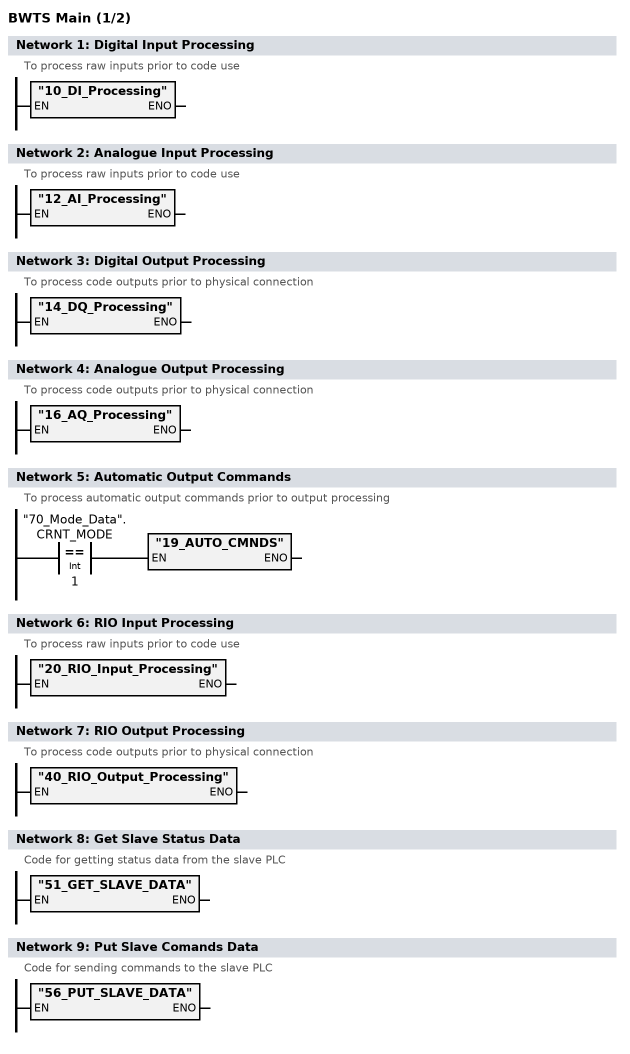
   RUNG wire#powerrail
      "10_DI_Processing"()
   END_RUNG
   // the same network as SCL:
   "10_DI_Processing"();
END_REGION

REGION Network 2: Analogue Input Processing
   // To process raw inputs prior to code use
   RUNG wire#powerrail
      "12_AI_Processing"()
   END_RUNG
   // the same network as SCL:
   "12_AI_Processing"();
END_REGION

REGION Network 3: Digital Output Processing
   // To process code outputs prior to physical connection
   RUNG wire#powerrail
      "14_DQ_Processing"()
   END_RUNG
   // the same network as SCL:
   "14_DQ_Processing"();
END_REGION

REGION Network 4: Analogue Output Processing
   // To process code outputs prior to physical connection
   RUNG wire#powerrail
      "16_AQ_Processing"()
   END_RUNG
   // the same network as SCL:
   "16_AQ_Processing"();
END_REGION

REGION Network 5: Automatic Output Commands
   // To process automatic output commands prior to output processing
   RUNG wire#powerrail
      { S7_Templates := "SrcType := Int" } EQ_Contact(in1 := "70_Mode_Data".CRNT_MODE, in2 := 1)
      "19_AUTO_CMNDS"()
   END_RUNG
   // the same network as SCL:
   IF "70_Mode_Data".CRNT_MODE = 1 THEN "19_AUTO_CMNDS"(); END_IF;
END_REGION

REGION Network 6: RIO Input Processing
   // To process raw inputs prior to code use
   RUNG wire#powerrail
      "20_RIO_Input_Processing"()
   END_RUNG
   // the same network as SCL:
   "20_RIO_Input_Processing"();
END_REGION

REGION Network 7: RIO Output Processing
   // To process code outputs prior to physical connection
   RUNG wire#powerrail
      "40_RIO_Output_Processing"()
   END_RUNG
   // the same network as SCL:
   "40_RIO_Output_Processing"();
END_REGION

REGION Network 8: Get Slave Status Data
   // Code for getting status data from the slave PLC
   RUNG wire#powerrail
      "51_GET_SLAVE_DATA"()
   END_RUNG
   // the same network as SCL:
   "51_GET_SLAVE_DATA"();
END_REGION

REGION Network 9: Put Slave Comands Data
   // Code for sending commands to the slave PLC
   RUNG wire#powerrail
      "56_PUT_SLAVE_DATA"()
   END_RUNG
   // the same network as SCL:
   "56_PUT_SLAVE_DATA"();
END_REGION

REGION Network 10: Communications Heart Beat
   // Code for communications heart beat bit
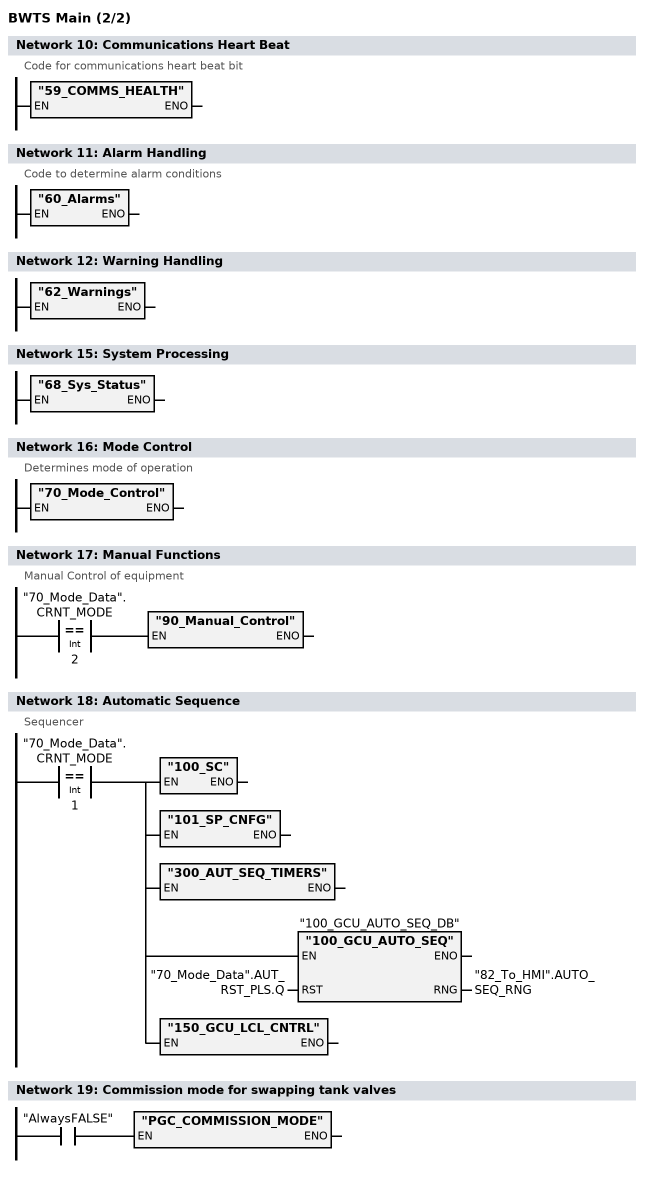
   RUNG wire#powerrail
      "59_COMMS_HEALTH"()
   END_RUNG
   // the same network as SCL:
   "59_COMMS_HEALTH"();
END_REGION

REGION Network 11: Alarm Handling
   // Code to determine alarm conditions
   RUNG wire#powerrail
      "60_Alarms"()
   END_RUNG
   // the same network as SCL:
   "60_Alarms"();
END_REGION

REGION Network 12: Warning Handling
   RUNG wire#powerrail
      "62_Warnings"()
   END_RUNG
   // the same network as SCL:
   "62_Warnings"();
END_REGION

REGION Network 13: Message Handling
   // Handles messaging
END_REGION

REGION Network 14: Event Handling
   // Records event data
END_REGION

REGION Network 15: System Processing
   RUNG wire#powerrail
      "68_Sys_Status"()
   END_RUNG
   // the same network as SCL:
   "68_Sys_Status"();
END_REGION

REGION Network 16: Mode Control
   // Determines mode of operation
   RUNG wire#powerrail
      "70_Mode_Control"()
   END_RUNG
   // the same network as SCL:
   "70_Mode_Control"();
END_REGION

REGION Network 17: Manual Functions
   // Manual Control of equipment
   RUNG wire#powerrail
      { S7_Templates := "SrcType := Int" } EQ_Contact(in1 := "70_Mode_Data".CRNT_MODE, in2 := 2)
      "90_Manual_Control"()
   END_RUNG
   // the same network as SCL:
   IF "70_Mode_Data".CRNT_MODE = 2 THEN "90_Manual_Control"(); END_IF;
END_REGION

REGION Network 18: Automatic Sequence
   // Sequencer
   RUNG wire#powerrail
      { S7_Templates := "SrcType := Int" } EQ_Contact(in1 := "70_Mode_Data".CRNT_MODE, in2 := 1)
      wire#w1
      "100_SC"()
   END_RUNG
   RUNG wire#w1
      "101_SP_CNFG"()
   END_RUNG
   RUNG wire#w1
      "300_AUT_SEQ_TIMERS"()
   END_RUNG
   RUNG wire#w1
      "100_GCU_AUTO_SEQ_DB"(RST := "70_Mode_Data".AUT_RST_PLS.Q, RNG => "82_To_HMI".AUTO_SEQ_RNG)
   END_RUNG
   RUNG wire#w1
      "150_GCU_LCL_CNTRL"()
   END_RUNG
   // the same network as SCL:
   #_w1 := "70_Mode_Data".CRNT_MODE = 1;
   IF #_w1 THEN
       "100_SC"();
       "101_SP_CNFG"();
       "300_AUT_SEQ_TIMERS"();
       "100_GCU_AUTO_SEQ_DB"(RST := "70_Mode_Data".AUT_RST_PLS.Q, RNG => "82_To_HMI".AUTO_SEQ_RNG);   // "100_GCU_AUTO_SEQ"
       "150_GCU_LCL_CNTRL"();
   END_IF;
END_REGION

REGION Network 19: Commission mode for swapping tank valves
   RUNG wire#powerrail
      Contact( "AlwaysFALSE" )
      "PGC_COMMISSION_MODE"()
   END_RUNG
   // the same network as SCL:
   IF "AlwaysFALSE" THEN "PGC_COMMISSION_MODE"(); END_IF;
END_REGION
END_ORGANIZATION_BLOCK

// folder: 10 - 19 IO & Processing

FUNCTION "10_DI_Processing" : Void   // FC10, LAD
TITLE = Digital Input Processing
{ S7_Optimized_Access := 'TRUE' }
AUTHOR : JRS
VERSION : 0.1
// To process raw inputs prior to code use
BEGIN

REGION Network 1: I136.0 - Spare Input
   // True = N/A, False = N/A
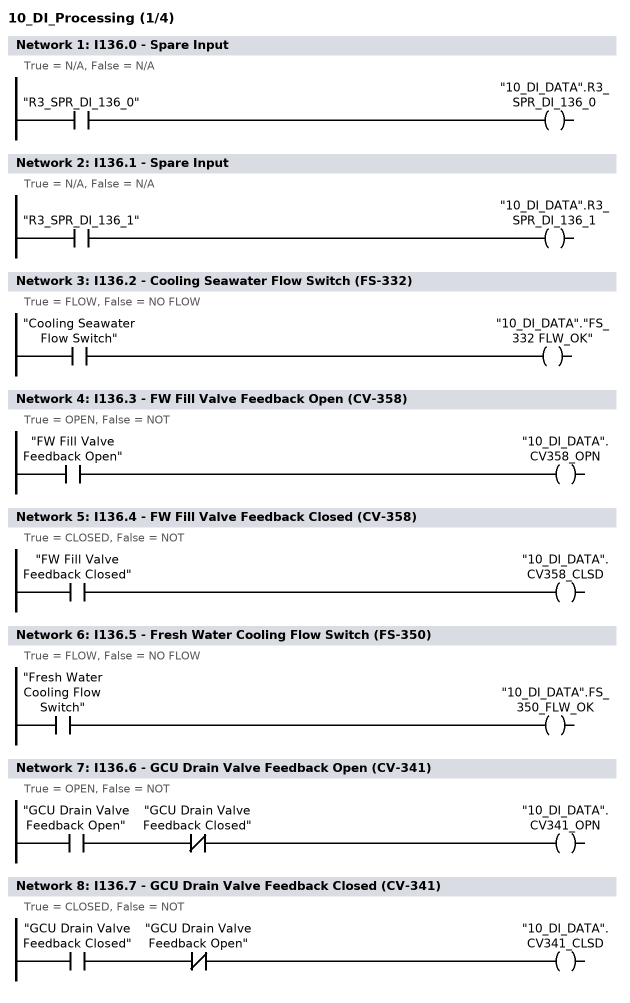
   RUNG wire#powerrail
      Contact( "R3_SPR_DI_136_0" )
      Coil( "10_DI_DATA".R3_SPR_DI_136_0 )
   END_RUNG
   // the same network as SCL:
   "10_DI_DATA".R3_SPR_DI_136_0 := "R3_SPR_DI_136_0";
END_REGION

REGION Network 2: I136.1 - Spare Input
   // True = N/A, False = N/A
   RUNG wire#powerrail
      Contact( "R3_SPR_DI_136_1" )
      Coil( "10_DI_DATA".R3_SPR_DI_136_1 )
   END_RUNG
   // the same network as SCL:
   "10_DI_DATA".R3_SPR_DI_136_1 := "R3_SPR_DI_136_1";
END_REGION

REGION Network 3: I136.2 - Cooling Seawater Flow Switch (FS-332)
   // True = FLOW, False = NO FLOW
   RUNG wire#powerrail
      Contact( "Cooling Seawater Flow Switch" )
      Coil( "10_DI_DATA"."FS_332 FLW_OK" )
   END_RUNG
   // the same network as SCL:
   "10_DI_DATA"."FS_332 FLW_OK" := "Cooling Seawater Flow Switch";
END_REGION

REGION Network 4: I136.3 - FW Fill Valve Feedback Open (CV-358)
   // True = OPEN, False = NOT
   RUNG wire#powerrail
      Contact( "FW Fill Valve Feedback Open" )
      Coil( "10_DI_DATA".CV358_OPN )
   END_RUNG
   // the same network as SCL:
   "10_DI_DATA".CV358_OPN := "FW Fill Valve Feedback Open";
END_REGION

REGION Network 5: I136.4 - FW Fill Valve Feedback Closed (CV-358)
   // True = CLOSED, False = NOT
   RUNG wire#powerrail
      Contact( "FW Fill Valve Feedback Closed" )
      Coil( "10_DI_DATA".CV358_CLSD )
   END_RUNG
   // the same network as SCL:
   "10_DI_DATA".CV358_CLSD := "FW Fill Valve Feedback Closed";
END_REGION

REGION Network 6: I136.5 - Fresh Water Cooling Flow Switch (FS-350)
   // True = FLOW, False = NO FLOW
   RUNG wire#powerrail
      Contact( "Fresh Water Cooling Flow Switch" )
      Coil( "10_DI_DATA".FS_350_FLW_OK )
   END_RUNG
   // the same network as SCL:
   "10_DI_DATA".FS_350_FLW_OK := "Fresh Water Cooling Flow Switch";
END_REGION

REGION Network 7: I136.6 - GCU Drain Valve Feedback Open (CV-341)
   // True = OPEN, False = NOT
   RUNG wire#powerrail
      Contact( "GCU Drain Valve Feedback Open" )
      I_Contact( "GCU Drain Valve Feedback Closed" )
      Coil( "10_DI_DATA".CV341_OPN )
   END_RUNG
   // the same network as SCL:
   "10_DI_DATA".CV341_OPN := "GCU Drain Valve Feedback Open" AND NOT "GCU Drain Valve Feedback Closed";
END_REGION

REGION Network 8: I136.7 - GCU Drain Valve Feedback Closed (CV-341)
   // True = CLOSED, False = NOT
   RUNG wire#powerrail
      Contact( "GCU Drain Valve Feedback Closed" )
      I_Contact( "GCU Drain Valve Feedback Open" )
      Coil( "10_DI_DATA".CV341_CLSD )
   END_RUNG
   // the same network as SCL:
   "10_DI_DATA".CV341_CLSD := "GCU Drain Valve Feedback Closed" AND NOT "GCU Drain Valve Feedback Open";
END_REGION

REGION Network 9: I137.0 - Gas to Deck Valve Feedback Open (CV-406)
   // True = OPEN, False = NOT
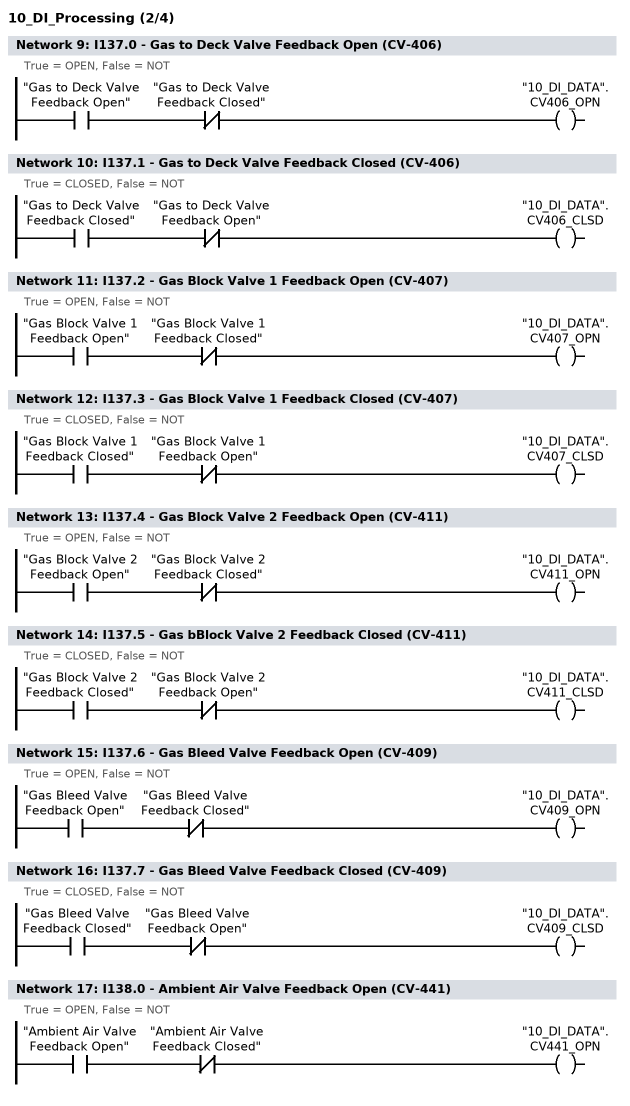
   RUNG wire#powerrail
      Contact( "Gas to Deck Valve Feedback Open" )
      I_Contact( "Gas to Deck Valve Feedback Closed" )
      Coil( "10_DI_DATA".CV406_OPN )
   END_RUNG
   // the same network as SCL:
   "10_DI_DATA".CV406_OPN := "Gas to Deck Valve Feedback Open" AND NOT "Gas to Deck Valve Feedback Closed";
END_REGION

REGION Network 10: I137.1 - Gas to Deck Valve Feedback Closed (CV-406)
   // True = CLOSED, False = NOT
   RUNG wire#powerrail
      Contact( "Gas to Deck Valve Feedback Closed" )
      I_Contact( "Gas to Deck Valve Feedback Open" )
      Coil( "10_DI_DATA".CV406_CLSD )
   END_RUNG
   // the same network as SCL:
   "10_DI_DATA".CV406_CLSD := "Gas to Deck Valve Feedback Closed" AND NOT "Gas to Deck Valve Feedback Open";
END_REGION

REGION Network 11: I137.2 - Gas Block Valve 1 Feedback Open (CV-407)
   // True = OPEN, False = NOT
   RUNG wire#powerrail
      Contact( "Gas Block Valve 1 Feedback Open" )
      I_Contact( "Gas Block Valve 1 Feedback Closed" )
      Coil( "10_DI_DATA".CV407_OPN )
   END_RUNG
   // the same network as SCL:
   "10_DI_DATA".CV407_OPN := "Gas Block Valve 1 Feedback Open" AND NOT "Gas Block Valve 1 Feedback Closed";
END_REGION

REGION Network 12: I137.3 - Gas Block Valve 1 Feedback Closed (CV-407)
   // True = CLOSED, False = NOT
   RUNG wire#powerrail
      Contact( "Gas Block Valve 1 Feedback Closed" )
      I_Contact( "Gas Block Valve 1 Feedback Open" )
      Coil( "10_DI_DATA".CV407_CLSD )
   END_RUNG
   // the same network as SCL:
   "10_DI_DATA".CV407_CLSD := "Gas Block Valve 1 Feedback Closed" AND NOT "Gas Block Valve 1 Feedback Open";
END_REGION

REGION Network 13: I137.4 - Gas Block Valve 2 Feedback Open (CV-411)
   // True = OPEN, False = NOT
   RUNG wire#powerrail
      Contact( "Gas Block Valve 2 Feedback Open" )
      I_Contact( "Gas Block Valve 2 Feedback Closed" )
      Coil( "10_DI_DATA".CV411_OPN )
   END_RUNG
   // the same network as SCL:
   "10_DI_DATA".CV411_OPN := "Gas Block Valve 2 Feedback Open" AND NOT "Gas Block Valve 2 Feedback Closed";
END_REGION

REGION Network 14: I137.5 - Gas bBlock Valve 2 Feedback Closed (CV-411)
   // True = CLOSED, False = NOT
   RUNG wire#powerrail
      Contact( "Gas Block Valve 2 Feedback Closed" )
      I_Contact( "Gas Block Valve 2 Feedback Open" )
      Coil( "10_DI_DATA".CV411_CLSD )
   END_RUNG
   // the same network as SCL:
   "10_DI_DATA".CV411_CLSD := "Gas Block Valve 2 Feedback Closed" AND NOT "Gas Block Valve 2 Feedback Open";
END_REGION

REGION Network 15: I137.6 - Gas Bleed Valve Feedback Open (CV-409)
   // True = OPEN, False = NOT
   RUNG wire#powerrail
      Contact( "Gas Bleed Valve Feedback Open" )
      I_Contact( "Gas Bleed Valve Feedback Closed" )
      Coil( "10_DI_DATA".CV409_OPN )
   END_RUNG
   // the same network as SCL:
   "10_DI_DATA".CV409_OPN := "Gas Bleed Valve Feedback Open" AND NOT "Gas Bleed Valve Feedback Closed";
END_REGION

REGION Network 16: I137.7 - Gas Bleed Valve Feedback Closed (CV-409)
   // True = CLOSED, False = NOT
   RUNG wire#powerrail
      Contact( "Gas Bleed Valve Feedback Closed" )
      I_Contact( "Gas Bleed Valve Feedback Open" )
      Coil( "10_DI_DATA".CV409_CLSD )
   END_RUNG
   // the same network as SCL:
   "10_DI_DATA".CV409_CLSD := "Gas Bleed Valve Feedback Closed" AND NOT "Gas Bleed Valve Feedback Open";
END_REGION

REGION Network 17: I138.0 - Ambient Air Valve Feedback Open (CV-441)
   // True = OPEN, False = NOT
   RUNG wire#powerrail
      Contact( "Ambient Air Valve Feedback Open" )
      I_Contact( "Ambient Air Valve Feedback Closed" )
      Coil( "10_DI_DATA".CV441_OPN )
   END_RUNG
   // the same network as SCL:
   "10_DI_DATA".CV441_OPN := "Ambient Air Valve Feedback Open" AND NOT "Ambient Air Valve Feedback Closed";
END_REGION

REGION Network 18: I138.1 - Ambient Air Valve Feedback Closed (CV-441)
   // True = CLOSED, False = NOT
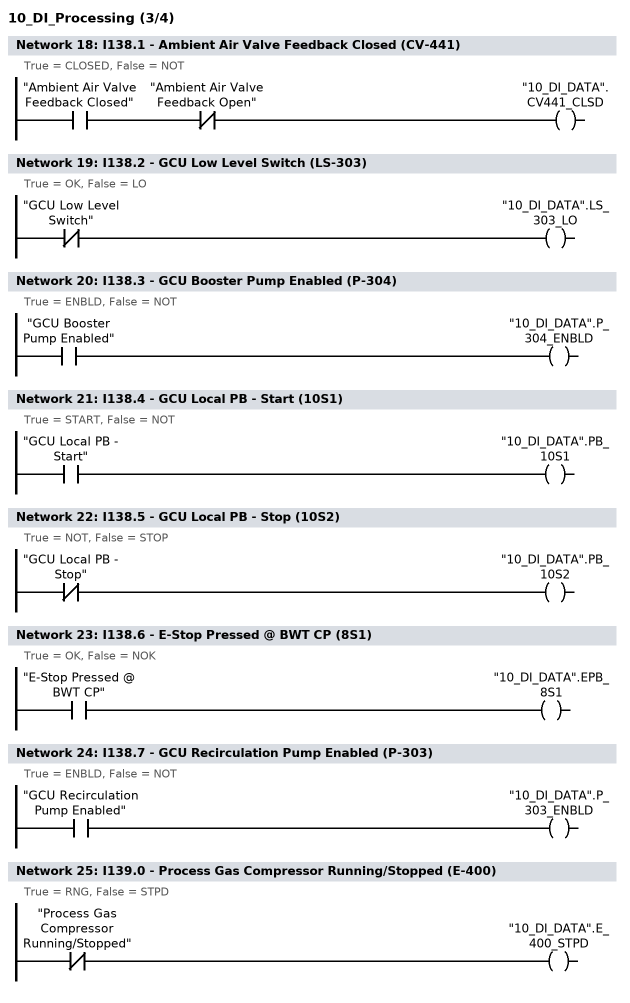
   RUNG wire#powerrail
      Contact( "Ambient Air Valve Feedback Closed" )
      I_Contact( "Ambient Air Valve Feedback Open" )
      Coil( "10_DI_DATA".CV441_CLSD )
   END_RUNG
   // the same network as SCL:
   "10_DI_DATA".CV441_CLSD := "Ambient Air Valve Feedback Closed" AND NOT "Ambient Air Valve Feedback Open";
END_REGION

REGION Network 19: I138.2 - GCU Low Level Switch (LS-303)
   // True = OK, False = LO
   RUNG wire#powerrail
      I_Contact( "GCU Low Level Switch" )
      Coil( "10_DI_DATA".LS_303_LO )
   END_RUNG
   // the same network as SCL:
   "10_DI_DATA".LS_303_LO := NOT "GCU Low Level Switch";
END_REGION

REGION Network 20: I138.3 - GCU Booster Pump Enabled (P-304)
   // True = ENBLD, False = NOT
   RUNG wire#powerrail
      Contact( "GCU Booster Pump Enabled" )
      Coil( "10_DI_DATA".P_304_ENBLD )
   END_RUNG
   // the same network as SCL:
   "10_DI_DATA".P_304_ENBLD := "GCU Booster Pump Enabled";
END_REGION

REGION Network 21: I138.4 - GCU Local PB - Start (10S1)
   // True = START, False = NOT
   RUNG wire#powerrail
      Contact( "GCU Local PB - Start" )
      Coil( "10_DI_DATA".PB_10S1 )
   END_RUNG
   // the same network as SCL:
   "10_DI_DATA".PB_10S1 := "GCU Local PB - Start";
END_REGION

REGION Network 22: I138.5 - GCU Local PB - Stop (10S2)
   // True = NOT, False = STOP
   RUNG wire#powerrail
      I_Contact( "GCU Local PB - Stop" )
      Coil( "10_DI_DATA".PB_10S2 )
   END_RUNG
   // the same network as SCL:
   "10_DI_DATA".PB_10S2 := NOT "GCU Local PB - Stop";
END_REGION

REGION Network 23: I138.6 - E-Stop Pressed @ BWT CP (8S1)
   // True = OK, False = NOK
   RUNG wire#powerrail
      Contact( "E-Stop Pressed @ BWT CP" )
      Coil( "10_DI_DATA".EPB_8S1 )
   END_RUNG
   // the same network as SCL:
   "10_DI_DATA".EPB_8S1 := "E-Stop Pressed @ BWT CP";
END_REGION

REGION Network 24: I138.7 - GCU Recirculation Pump Enabled (P-303)
   // True = ENBLD, False = NOT
   RUNG wire#powerrail
      Contact( "GCU Recirculation Pump Enabled" )
      Coil( "10_DI_DATA".P_303_ENBLD )
   END_RUNG
   // the same network as SCL:
   "10_DI_DATA".P_303_ENBLD := "GCU Recirculation Pump Enabled";
END_REGION

REGION Network 25: I139.0 - Process Gas Compressor Running/Stopped (E-400)
   // True = RNG, False = STPD
   RUNG wire#powerrail
      I_Contact( "Process Gas Compressor Running/Stopped" )
      Coil( "10_DI_DATA".E_400_STPD )
   END_RUNG
   // the same network as SCL:
   "10_DI_DATA".E_400_STPD := NOT "Process Gas Compressor Running/Stopped";
END_REGION

REGION Network 26: I139.1 - Process Gas Compressor Tripped/Shutdown (E-400)
   // True = NOK, False = OK
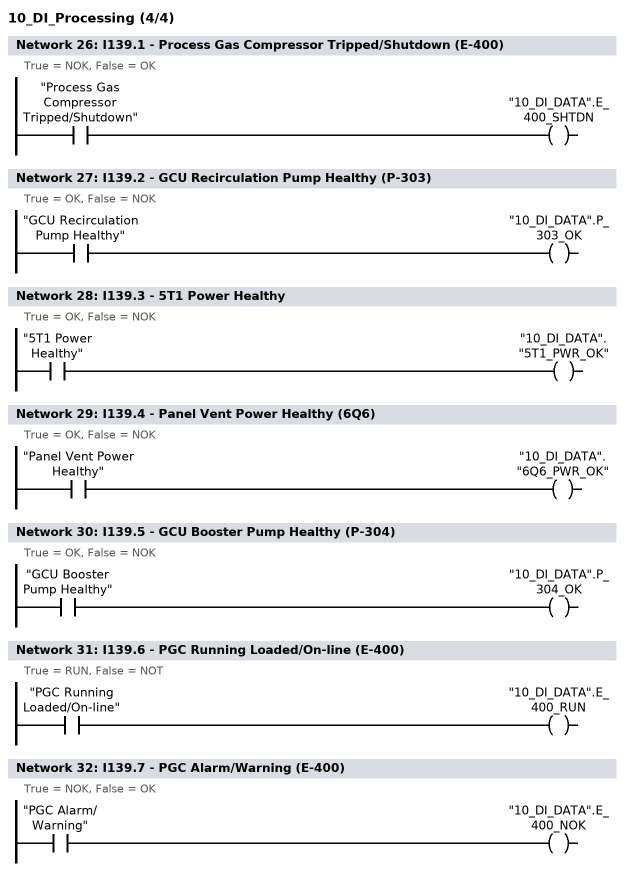
   RUNG wire#powerrail
      Contact( "Process Gas Compressor Tripped/Shutdown" )
      Coil( "10_DI_DATA".E_400_SHTDN )
   END_RUNG
   // the same network as SCL:
   "10_DI_DATA".E_400_SHTDN := "Process Gas Compressor Tripped/Shutdown";
END_REGION

REGION Network 27: I139.2 - GCU Recirculation Pump Healthy (P-303)
   // True = OK, False = NOK
   RUNG wire#powerrail
      Contact( "GCU Recirculation Pump Healthy" )
      Coil( "10_DI_DATA".P_303_OK )
   END_RUNG
   // the same network as SCL:
   "10_DI_DATA".P_303_OK := "GCU Recirculation Pump Healthy";
END_REGION

REGION Network 28: I139.3 - 5T1 Power Healthy
   // True = OK, False = NOK
   RUNG wire#powerrail
      Contact( "5T1 Power Healthy" )
      Coil( "10_DI_DATA"."5T1_PWR_OK" )
   END_RUNG
   // the same network as SCL:
   "10_DI_DATA"."5T1_PWR_OK" := "5T1 Power Healthy";
END_REGION

REGION Network 29: I139.4 - Panel Vent Power Healthy (6Q6)
   // True = OK, False = NOK
   RUNG wire#powerrail
      Contact( "Panel Vent Power Healthy" )
      Coil( "10_DI_DATA"."6Q6_PWR_OK" )
   END_RUNG
   // the same network as SCL:
   "10_DI_DATA"."6Q6_PWR_OK" := "Panel Vent Power Healthy";
END_REGION

REGION Network 30: I139.5 - GCU Booster Pump Healthy (P-304)
   // True = OK, False = NOK
   RUNG wire#powerrail
      Contact( "GCU Booster Pump Healthy" )
      Coil( "10_DI_DATA".P_304_OK )
   END_RUNG
   // the same network as SCL:
   "10_DI_DATA".P_304_OK := "GCU Booster Pump Healthy";
END_REGION

REGION Network 31: I139.6 - PGC Running Loaded/On-line (E-400)
   // True = RUN, False = NOT
   RUNG wire#powerrail
      Contact( "PGC Running Loaded/On-line" )
      Coil( "10_DI_DATA".E_400_RUN )
   END_RUNG
   // the same network as SCL:
   "10_DI_DATA".E_400_RUN := "PGC Running Loaded/On-line";
END_REGION

REGION Network 32: I139.7 - PGC Alarm/Warning (E-400)
   // True = NOK, False = OK
   RUNG wire#powerrail
      Contact( "PGC Alarm/Warning" )
      Coil( "10_DI_DATA".E_400_NOK )
   END_RUNG
   // the same network as SCL:
   "10_DI_DATA".E_400_NOK := "PGC Alarm/Warning";
END_REGION
END_FUNCTION

FUNCTION "12_AI_Processing" : Void   // FC12, LAD
TITLE = Analogue Input Processing
{ S7_Optimized_Access := 'TRUE' }
AUTHOR : JRS
VERSION : 0.1
// To process raw inputs prior to code use
BEGIN

REGION Network 1: IW800 - GCU Level (LIT-304)
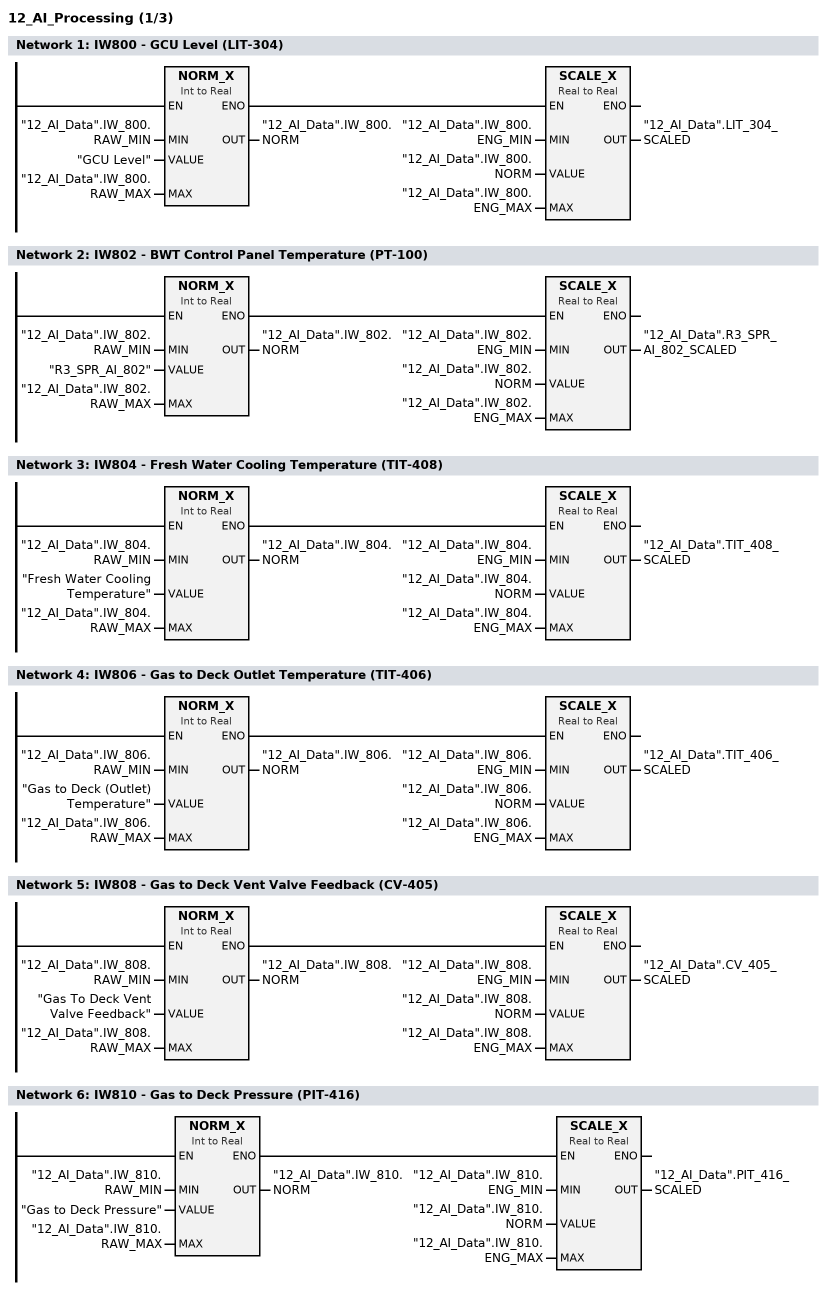
   RUNG wire#powerrail
      { S7_Templates := "[SrcType := Int, DestType := Real]" } Normalize(min := "12_AI_Data".IW_800.RAW_MIN, value := "GCU Level", max := "12_AI_Data".IW_800.RAW_MAX, out => "12_AI_Data".IW_800.NORM)
      { S7_Templates := "[SrcType := Real, DestType := Real]" } Scale(min := "12_AI_Data".IW_800.ENG_MIN, value := "12_AI_Data".IW_800.NORM, max := "12_AI_Data".IW_800.ENG_MAX, out => "12_AI_Data".LIT_304_SCALED)
   END_RUNG
   // the same network as SCL:
   "12_AI_Data".IW_800.NORM := NORM_X(MIN := "12_AI_Data".IW_800.RAW_MIN, VALUE := "GCU Level", MAX := "12_AI_Data".IW_800.RAW_MAX);
   "12_AI_Data".LIT_304_SCALED := SCALE_X(MIN := "12_AI_Data".IW_800.ENG_MIN, VALUE := "12_AI_Data".IW_800.NORM, MAX := "12_AI_Data".IW_800.ENG_MAX);
END_REGION

REGION Network 2: IW802 - BWT Control Panel Temperature (PT-100)
   RUNG wire#powerrail
      { S7_Templates := "[SrcType := Int, DestType := Real]" } Normalize(min := "12_AI_Data".IW_802.RAW_MIN, value := "R3_SPR_AI_802", max := "12_AI_Data".IW_802.RAW_MAX, out => "12_AI_Data".IW_802.NORM)
      { S7_Templates := "[SrcType := Real, DestType := Real]" } Scale(min := "12_AI_Data".IW_802.ENG_MIN, value := "12_AI_Data".IW_802.NORM, max := "12_AI_Data".IW_802.ENG_MAX, out => "12_AI_Data".R3_SPR_AI_802_SCALED)
   END_RUNG
   // the same network as SCL:
   "12_AI_Data".IW_802.NORM := NORM_X(MIN := "12_AI_Data".IW_802.RAW_MIN, VALUE := "R3_SPR_AI_802", MAX := "12_AI_Data".IW_802.RAW_MAX);
   "12_AI_Data".R3_SPR_AI_802_SCALED := SCALE_X(MIN := "12_AI_Data".IW_802.ENG_MIN, VALUE := "12_AI_Data".IW_802.NORM, MAX := "12_AI_Data".IW_802.ENG_MAX);
END_REGION

REGION Network 3: IW804 - Fresh Water Cooling Temperature (TIT-408)
   RUNG wire#powerrail
      { S7_Templates := "[SrcType := Int, DestType := Real]" } Normalize(min := "12_AI_Data".IW_804.RAW_MIN, value := "Fresh Water Cooling Temperature", max := "12_AI_Data".IW_804.RAW_MAX, out => "12_AI_Data".IW_804.NORM)
      { S7_Templates := "[SrcType := Real, DestType := Real]" } Scale(min := "12_AI_Data".IW_804.ENG_MIN, value := "12_AI_Data".IW_804.NORM, max := "12_AI_Data".IW_804.ENG_MAX, out => "12_AI_Data".TIT_408_SCALED)
   END_RUNG
   // the same network as SCL:
   "12_AI_Data".IW_804.NORM := NORM_X(MIN := "12_AI_Data".IW_804.RAW_MIN, VALUE := "Fresh Water Cooling Temperature", MAX := "12_AI_Data".IW_804.RAW_MAX);
   "12_AI_Data".TIT_408_SCALED := SCALE_X(MIN := "12_AI_Data".IW_804.ENG_MIN, VALUE := "12_AI_Data".IW_804.NORM, MAX := "12_AI_Data".IW_804.ENG_MAX);
END_REGION

REGION Network 4: IW806 - Gas to Deck Outlet Temperature (TIT-406)
   RUNG wire#powerrail
      { S7_Templates := "[SrcType := Int, DestType := Real]" } Normalize(min := "12_AI_Data".IW_806.RAW_MIN, value := "Gas to Deck (Outlet) Temperature", max := "12_AI_Data".IW_806.RAW_MAX, out => "12_AI_Data".IW_806.NORM)
      { S7_Templates := "[SrcType := Real, DestType := Real]" } Scale(min := "12_AI_Data".IW_806.ENG_MIN, value := "12_AI_Data".IW_806.NORM, max := "12_AI_Data".IW_806.ENG_MAX, out => "12_AI_Data".TIT_406_SCALED)
   END_RUNG
   // the same network as SCL:
   "12_AI_Data".IW_806.NORM := NORM_X(MIN := "12_AI_Data".IW_806.RAW_MIN, VALUE := "Gas to Deck (Outlet) Temperature", MAX := "12_AI_Data".IW_806.RAW_MAX);
   "12_AI_Data".TIT_406_SCALED := SCALE_X(MIN := "12_AI_Data".IW_806.ENG_MIN, VALUE := "12_AI_Data".IW_806.NORM, MAX := "12_AI_Data".IW_806.ENG_MAX);
END_REGION

REGION Network 5: IW808 - Gas to Deck Vent Valve Feedback (CV-405)
   RUNG wire#powerrail
      { S7_Templates := "[SrcType := Int, DestType := Real]" } Normalize(min := "12_AI_Data".IW_808.RAW_MIN, value := "Gas To Deck Vent Valve Feedback", max := "12_AI_Data".IW_808.RAW_MAX, out => "12_AI_Data".IW_808.NORM)
      { S7_Templates := "[SrcType := Real, DestType := Real]" } Scale(min := "12_AI_Data".IW_808.ENG_MIN, value := "12_AI_Data".IW_808.NORM, max := "12_AI_Data".IW_808.ENG_MAX, out => "12_AI_Data".CV_405_SCALED)
   END_RUNG
   // the same network as SCL:
   "12_AI_Data".IW_808.NORM := NORM_X(MIN := "12_AI_Data".IW_808.RAW_MIN, VALUE := "Gas To Deck Vent Valve Feedback", MAX := "12_AI_Data".IW_808.RAW_MAX);
   "12_AI_Data".CV_405_SCALED := SCALE_X(MIN := "12_AI_Data".IW_808.ENG_MIN, VALUE := "12_AI_Data".IW_808.NORM, MAX := "12_AI_Data".IW_808.ENG_MAX);
END_REGION

REGION Network 6: IW810 - Gas to Deck Pressure (PIT-416)
   RUNG wire#powerrail
      { S7_Templates := "[SrcType := Int, DestType := Real]" } Normalize(min := "12_AI_Data".IW_810.RAW_MIN, value := "Gas to Deck Pressure", max := "12_AI_Data".IW_810.RAW_MAX, out => "12_AI_Data".IW_810.NORM)
      { S7_Templates := "[SrcType := Real, DestType := Real]" } Scale(min := "12_AI_Data".IW_810.ENG_MIN, value := "12_AI_Data".IW_810.NORM, max := "12_AI_Data".IW_810.ENG_MAX, out => "12_AI_Data".PIT_416_SCALED)
   END_RUNG
   // the same network as SCL:
   "12_AI_Data".IW_810.NORM := NORM_X(MIN := "12_AI_Data".IW_810.RAW_MIN, VALUE := "Gas to Deck Pressure", MAX := "12_AI_Data".IW_810.RAW_MAX);
   "12_AI_Data".PIT_416_SCALED := SCALE_X(MIN := "12_AI_Data".IW_810.ENG_MIN, VALUE := "12_AI_Data".IW_810.NORM, MAX := "12_AI_Data".IW_810.ENG_MAX);
END_REGION

REGION Network 7: IW812 - Fresh Water Inlet Pressure (PIT-358)
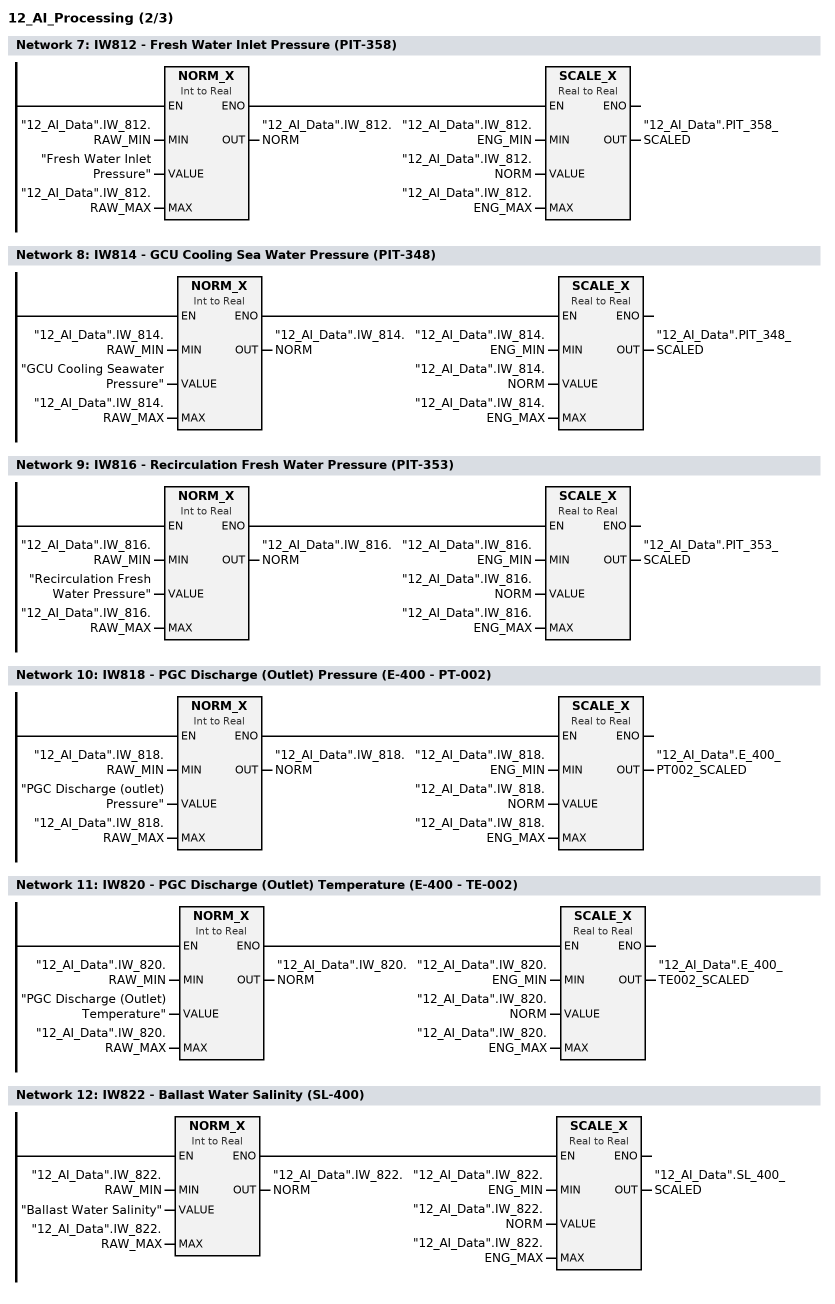
   RUNG wire#powerrail
      { S7_Templates := "[SrcType := Int, DestType := Real]" } Normalize(min := "12_AI_Data".IW_812.RAW_MIN, value := "Fresh Water Inlet Pressure", max := "12_AI_Data".IW_812.RAW_MAX, out => "12_AI_Data".IW_812.NORM)
      { S7_Templates := "[SrcType := Real, DestType := Real]" } Scale(min := "12_AI_Data".IW_812.ENG_MIN, value := "12_AI_Data".IW_812.NORM, max := "12_AI_Data".IW_812.ENG_MAX, out => "12_AI_Data".PIT_358_SCALED)
   END_RUNG
   // the same network as SCL:
   "12_AI_Data".IW_812.NORM := NORM_X(MIN := "12_AI_Data".IW_812.RAW_MIN, VALUE := "Fresh Water Inlet Pressure", MAX := "12_AI_Data".IW_812.RAW_MAX);
   "12_AI_Data".PIT_358_SCALED := SCALE_X(MIN := "12_AI_Data".IW_812.ENG_MIN, VALUE := "12_AI_Data".IW_812.NORM, MAX := "12_AI_Data".IW_812.ENG_MAX);
END_REGION

REGION Network 8: IW814 - GCU Cooling Sea Water Pressure (PIT-348)
   RUNG wire#powerrail
      { S7_Templates := "[SrcType := Int, DestType := Real]" } Normalize(min := "12_AI_Data".IW_814.RAW_MIN, value := "GCU Cooling Seawater Pressure", max := "12_AI_Data".IW_814.RAW_MAX, out => "12_AI_Data".IW_814.NORM)
      { S7_Templates := "[SrcType := Real, DestType := Real]" } Scale(min := "12_AI_Data".IW_814.ENG_MIN, value := "12_AI_Data".IW_814.NORM, max := "12_AI_Data".IW_814.ENG_MAX, out => "12_AI_Data".PIT_348_SCALED)
   END_RUNG
   // the same network as SCL:
   "12_AI_Data".IW_814.NORM := NORM_X(MIN := "12_AI_Data".IW_814.RAW_MIN, VALUE := "GCU Cooling Seawater Pressure", MAX := "12_AI_Data".IW_814.RAW_MAX);
   "12_AI_Data".PIT_348_SCALED := SCALE_X(MIN := "12_AI_Data".IW_814.ENG_MIN, VALUE := "12_AI_Data".IW_814.NORM, MAX := "12_AI_Data".IW_814.ENG_MAX);
END_REGION

REGION Network 9: IW816 - Recirculation Fresh Water Pressure (PIT-353)
   RUNG wire#powerrail
      { S7_Templates := "[SrcType := Int, DestType := Real]" } Normalize(min := "12_AI_Data".IW_816.RAW_MIN, value := "Recirculation Fresh Water Pressure", max := "12_AI_Data".IW_816.RAW_MAX, out => "12_AI_Data".IW_816.NORM)
      { S7_Templates := "[SrcType := Real, DestType := Real]" } Scale(min := "12_AI_Data".IW_816.ENG_MIN, value := "12_AI_Data".IW_816.NORM, max := "12_AI_Data".IW_816.ENG_MAX, out => "12_AI_Data".PIT_353_SCALED)
   END_RUNG
   // the same network as SCL:
   "12_AI_Data".IW_816.NORM := NORM_X(MIN := "12_AI_Data".IW_816.RAW_MIN, VALUE := "Recirculation Fresh Water Pressure", MAX := "12_AI_Data".IW_816.RAW_MAX);
   "12_AI_Data".PIT_353_SCALED := SCALE_X(MIN := "12_AI_Data".IW_816.ENG_MIN, VALUE := "12_AI_Data".IW_816.NORM, MAX := "12_AI_Data".IW_816.ENG_MAX);
END_REGION

REGION Network 10: IW818 - PGC Discharge (Outlet) Pressure (E-400 - PT-002)
   RUNG wire#powerrail
      { S7_Templates := "[SrcType := Int, DestType := Real]" } Normalize(min := "12_AI_Data".IW_818.RAW_MIN, value := "PGC Discharge (outlet) Pressure", max := "12_AI_Data".IW_818.RAW_MAX, out => "12_AI_Data".IW_818.NORM)
      { S7_Templates := "[SrcType := Real, DestType := Real]" } Scale(min := "12_AI_Data".IW_818.ENG_MIN, value := "12_AI_Data".IW_818.NORM, max := "12_AI_Data".IW_818.ENG_MAX, out => "12_AI_Data".E_400_PT002_SCALED)
   END_RUNG
   // the same network as SCL:
   "12_AI_Data".IW_818.NORM := NORM_X(MIN := "12_AI_Data".IW_818.RAW_MIN, VALUE := "PGC Discharge (outlet) Pressure", MAX := "12_AI_Data".IW_818.RAW_MAX);
   "12_AI_Data".E_400_PT002_SCALED := SCALE_X(MIN := "12_AI_Data".IW_818.ENG_MIN, VALUE := "12_AI_Data".IW_818.NORM, MAX := "12_AI_Data".IW_818.ENG_MAX);
END_REGION

REGION Network 11: IW820 - PGC Discharge (Outlet) Temperature (E-400 - TE-002)
   RUNG wire#powerrail
      { S7_Templates := "[SrcType := Int, DestType := Real]" } Normalize(min := "12_AI_Data".IW_820.RAW_MIN, value := "PGC Discharge (Outlet) Temperature", max := "12_AI_Data".IW_820.RAW_MAX, out => "12_AI_Data".IW_820.NORM)
      { S7_Templates := "[SrcType := Real, DestType := Real]" } Scale(min := "12_AI_Data".IW_820.ENG_MIN, value := "12_AI_Data".IW_820.NORM, max := "12_AI_Data".IW_820.ENG_MAX, out => "12_AI_Data".E_400_TE002_SCALED)
   END_RUNG
   // the same network as SCL:
   "12_AI_Data".IW_820.NORM := NORM_X(MIN := "12_AI_Data".IW_820.RAW_MIN, VALUE := "PGC Discharge (Outlet) Temperature", MAX := "12_AI_Data".IW_820.RAW_MAX);
   "12_AI_Data".E_400_TE002_SCALED := SCALE_X(MIN := "12_AI_Data".IW_820.ENG_MIN, VALUE := "12_AI_Data".IW_820.NORM, MAX := "12_AI_Data".IW_820.ENG_MAX);
END_REGION

REGION Network 12: IW822 - Ballast Water Salinity (SL-400)
   RUNG wire#powerrail
      { S7_Templates := "[SrcType := Int, DestType := Real]" } Normalize(min := "12_AI_Data".IW_822.RAW_MIN, value := "Ballast Water Salinity", max := "12_AI_Data".IW_822.RAW_MAX, out => "12_AI_Data".IW_822.NORM)
      { S7_Templates := "[SrcType := Real, DestType := Real]" } Scale(min := "12_AI_Data".IW_822.ENG_MIN, value := "12_AI_Data".IW_822.NORM, max := "12_AI_Data".IW_822.ENG_MAX, out => "12_AI_Data".SL_400_SCALED)
   END_RUNG
   // the same network as SCL:
   "12_AI_Data".IW_822.NORM := NORM_X(MIN := "12_AI_Data".IW_822.RAW_MIN, VALUE := "Ballast Water Salinity", MAX := "12_AI_Data".IW_822.RAW_MAX);
   "12_AI_Data".SL_400_SCALED := SCALE_X(MIN := "12_AI_Data".IW_822.ENG_MIN, VALUE := "12_AI_Data".IW_822.NORM, MAX := "12_AI_Data".IW_822.ENG_MAX);
END_REGION

